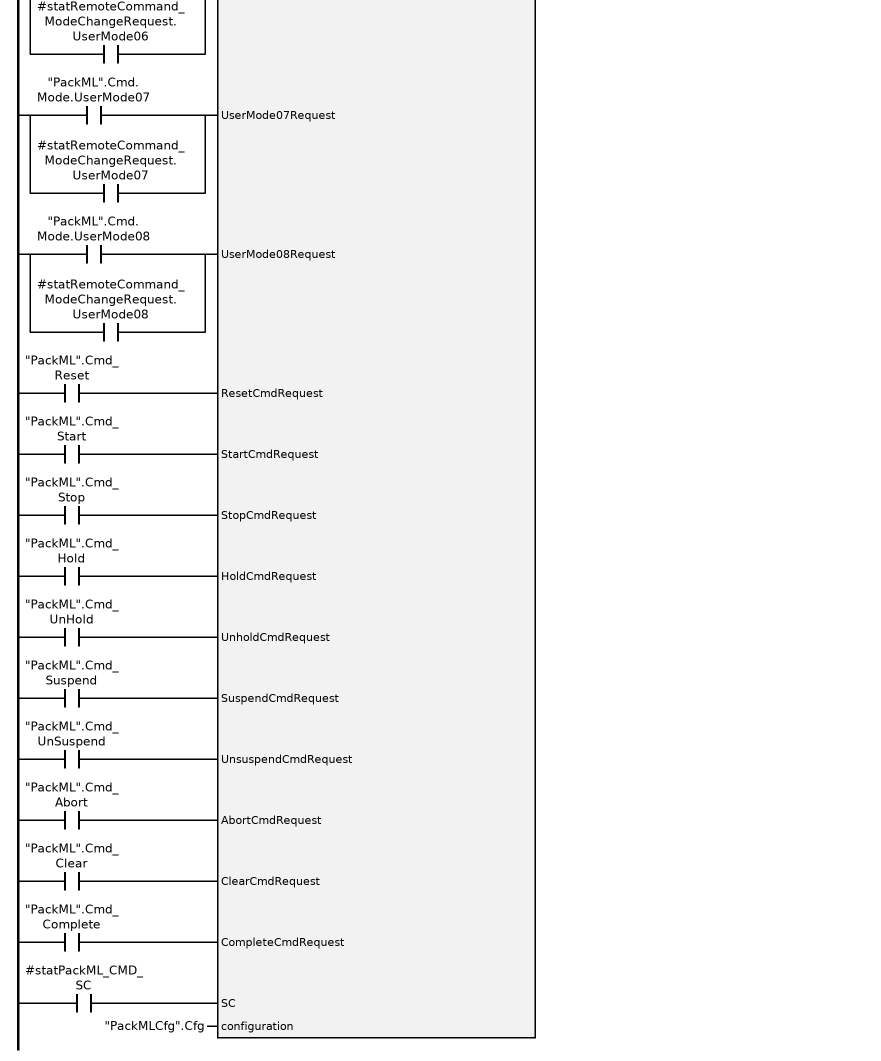
   RUNG wire#powerrail
      I_Contact( "FirstScan" )
      #instUnitModeStateManager(ProductionModeRequest := wire#w1, MaintenanceModeRequest := wire#w2, ManualModeRequest := wire#w3, UserMode01Request := wire#w4, UserMode02Request := wire#w5, UserMode03Request := wire#w6, UserMode04Request := wire#w7, UserMode05Request := wire#w8, UserMode06Request := wire#w9, UserMode07Request := wire#w10, UserMode08Request := wire#w11, ResetCmdRequest := wire#w12, StartCmdRequest := wire#w13, StopCmdRequest := wire#w14, HoldCmdRequest := wire#w15, UnholdCmdRequest := wire#w16, SuspendCmdRequest := wire#w17, UnsuspendCmdRequest := wire#w18, AbortCmdRequest := wire#w19, ClearCmdRequest := wire#w20, CompleteCmdRequest := wire#w21, SC := wire#w22, UnitMode :=, UnitModeChangeRequest := FALSE, CntrlCmd :=, CmdChangeRequest := FALSE, enableBooleanInterface := TRUE, configuration := "PackMLCfg".Cfg, UnitModeCurrent => "PackTags".Status.UnitModeCurrent, UnitModeRequested =>, UnitModeChangeInProcess => "PackTags".Status.UnitModeChangeInProcess, StateCurrent => "PackTags".Status.StateCurrent, StateRequested =>, StateChangeInProcess => "PackTags".Status.StateChangeInProcess, ProductionModeActive => "PackML".Sts.Mode.Production, MaintenanceModeActive => "PackML".Sts.Mode.Maintenance, ManualModeActive => "PackML".Sts.Mode.Manual, UserMode01Active => "PackML".Sts.Mode.UserMode01, UserMode02Active => "PackML".Sts.Mode.UserMode02, UserMode03Active => "PackML".Sts.Mode.UserMode03, UserMode04Active => "PackML".Sts.Mode.UserMode04, UserMode05Active => "PackML".Sts.Mode.UserMode05, UserMode06Active => "PackML".Sts.Mode.UserMode06, UserMode07Active => "PackML".Sts.Mode.UserMode07, UserMode08Active => "PackML".Sts.Mode.UserMode08, ClearingStateActive => "PackML".Sts.State.Clearing, StoppedStateActive => "PackML".Sts.State.Stopped, StartingStateActive => "PackML".Sts.State.Starting, IdleStateActive => "PackML".Sts.State.Idle, SuspendedStateActive => "PackML".Sts.State.Suspended, ExecuteStateActive => "PackML".Sts.State.Execute, StoppingStateActive => "PackML".Sts.State.Stopping, AbortingStateActive => "PackML".Sts.State.Aborting, AbortedStateActive => "PackML".Sts.State.Aborted, HoldingStateActive => "PackML".Sts.State.Holding, HeldStateActive => "PackML".Sts.State.Held, UnholdingStateActive => "PackML".Sts.State.Unholding, SuspendingStateActive => "PackML".Sts.State.Suspending, UnsuspendingStateActive => "PackML".Sts.State.Unsuspending, ResettingStateActive => "PackML".Sts.State.Resetting, CompletingStateActive => "PackML".Sts.State.Completing, CompleteStateActive => "PackML".Sts.State.Complete, StatesDisabled => "PackTags".Admin.StatesDisabled, diagnostics => "PackML".PackMLDiag)
      R_Coil( #statPackML_CMD_SC )
   END_RUNG
   RUNG wire#powerrail
      Contact( "PackML".Cmd.Mode.Production )
   END_RUNG wire#w1
   RUNG wire#powerrail
      Contact( #statRemoteCommand_ModeChangeRequest.Production )
   END_RUNG wire#w1
   RUNG wire#powerrail
      Contact( "PackML".Cmd.Mode.Maintenance )
   END_RUNG wire#w2
   RUNG wire#powerrail
      Contact( #statRemoteCommand_ModeChangeRequest.Maintenance )
   END_RUNG wire#w2
   RUNG wire#powerrail
      Contact( "PackML".Cmd.Mode.Manual )
   END_RUNG wire#w3
   RUNG wire#powerrail
      Contact( #statRemoteCommand_ModeChangeRequest.Manual )
   END_RUNG wire#w3
   RUNG wire#powerrail
      Contact( "PackML".Cmd.Mode.UserMode01 )
   END_RUNG wire#w4
   RUNG wire#powerrail
      Contact( #statRemoteCommand_ModeChangeRequest.UserMode01 )
   END_RUNG wire#w4
   RUNG wire#powerrail
      Contact( "PackML".Cmd.Mode.UserMode02 )
   END_RUNG wire#w5
   RUNG wire#powerrail
      Contact( #statRemoteCommand_ModeChangeRequest.UserMode02 )
   END_RUNG wire#w5
   RUNG wire#powerrail
      Contact( "PackML".Cmd.Mode.UserMode03 )
   END_RUNG wire#w6
   RUNG wire#powerrail
      Contact( #statRemoteCommand_ModeChangeRequest.UserMode03 )
   END_RUNG wire#w6
   RUNG wire#powerrail
      Contact( "PackML".Cmd.Mode.UserMode04 )
   END_RUNG wire#w7
   RUNG wire#powerrail
      Contact( #statRemoteCommand_ModeChangeRequest.UserMode04 )
   END_RUNG wire#w7
   RUNG wire#powerrail
      Contact( "PackML".Cmd.Mode.UserMode05 )
   END_RUNG wire#w8
   RUNG wire#powerrail
      Contact( #statRemoteCommand_ModeChangeRequest.UserMode05 )
   END_RUNG wire#w8
   RUNG wire#powerrail
      Contact( "PackML".Cmd.Mode.UserMode06 )
   END_RUNG wire#w9
   RUNG wire#powerrail
      Contact( #statRemoteCommand_ModeChangeRequest.UserMode06 )
   END_RUNG wire#w9
   RUNG wire#powerrail
      Contact( "PackML".Cmd.Mode.UserMode07 )
   END_RUNG wire#w10
   RUNG wire#powerrail
      Contact( #statRemoteCommand_ModeChangeRequest.UserMode07 )
   END_RUNG wire#w10
   RUNG wire#powerrail
      Contact( "PackML".Cmd.Mode.UserMode08 )
   END_RUNG wire#w11
   RUNG wire#powerrail
      Contact( #statRemoteCommand_ModeChangeRequest.UserMode08 )
   END_RUNG wire#w11
   RUNG wire#powerrail
      Contact( "PackML".Cmd_Reset )
   END_RUNG wire#w12
   RUNG wire#powerrail
      Contact( "PackML".Cmd_Start )
   END_RUNG wire#w13
   RUNG wire#powerrail
      Contact( "PackML".Cmd_Stop )
   END_RUNG wire#w14
   RUNG wire#powerrail
      Contact( "PackML".Cmd_Hold )
   END_RUNG wire#w15
   RUNG wire#powerrail
      Contact( "PackML".Cmd_UnHold )
   END_RUNG wire#w16
   RUNG wire#powerrail
      Contact( "PackML".Cmd_Suspend )
   END_RUNG wire#w17
   RUNG wire#powerrail
      Contact( "PackML".Cmd_UnSuspend )
   END_RUNG wire#w18
   RUNG wire#powerrail
      Contact( "PackML".Cmd_Abort )
   END_RUNG wire#w19
   RUNG wire#powerrail
      Contact( "PackML".Cmd_Clear )
   END_RUNG wire#w20
   RUNG wire#powerrail
      Contact( "PackML".Cmd_Complete )
   END_RUNG wire#w21
   RUNG wire#powerrail
      Contact( #statPackML_CMD_SC )
   END_RUNG wire#w22
   // the same network as SCL:
   #instUnitModeStateManager(EN := NOT "FirstScan",   // "LPMLV30_UnitModeStateManager"
                           UnitModeChangeRequest := FALSE,
                           CmdChangeRequest := FALSE,
                           enableBooleanInterface := TRUE,
                           ProductionModeRequest := "PackML".Cmd.Mode.Production OR #statRemoteCommand_ModeChangeRequest.Production,
                           MaintenanceModeRequest := "PackML".Cmd.Mode.Maintenance OR #statRemoteCommand_ModeChangeRequest.Maintenance,
                           ManualModeRequest := "PackML".Cmd.Mode.Manual OR #statRemoteCommand_ModeChangeRequest.Manual,
                           UserMode01Request := "PackML".Cmd.Mode.UserMode01 OR #statRemoteCommand_ModeChangeRequest.UserMode01,
                           UserMode02Request := "PackML".Cmd.Mode.UserMode02 OR #statRemoteCommand_ModeChangeRequest.UserMode02,
                           UserMode03Request := "PackML".Cmd.Mode.UserMode03 OR #statRemoteCommand_ModeChangeRequest.UserMode03,
                           UserMode04Request := "PackML".Cmd.Mode.UserMode04 OR #statRemoteCommand_ModeChangeRequest.UserMode04,
                           UserMode05Request := "PackML".Cmd.Mode.UserMode05 OR #statRemoteCommand_ModeChangeRequest.UserMode05,
                           UserMode06Request := "PackML".Cmd.Mode.UserMode06 OR #statRemoteCommand_ModeChangeRequest.UserMode06,
                           UserMode07Request := "PackML".Cmd.Mode.UserMode07 OR #statRemoteCommand_ModeChangeRequest.UserMode07,
                           UserMode08Request := "PackML".Cmd.Mode.UserMode08 OR #statRemoteCommand_ModeChangeRequest.UserMode08,
                           ResetCmdRequest := "PackML".Cmd_Reset,
                           StartCmdRequest := "PackML".Cmd_Start,
                           StopCmdRequest := "PackML".Cmd_Stop,
                           HoldCmdRequest := "PackML".Cmd_Hold,
                           UnholdCmdRequest := "PackML".Cmd_UnHold,
                           SuspendCmdRequest := "PackML".Cmd_Suspend,
                           UnsuspendCmdRequest := "PackML".Cmd_UnSuspend,
                           AbortCmdRequest := "PackML".Cmd_Abort,
                           ClearCmdRequest := "PackML".Cmd_Clear,
                           CompleteCmdRequest := "PackML".Cmd_Complete,
                           SC := #statPackML_CMD_SC,
                           configuration := "PackMLCfg".Cfg,
                           UnitModeCurrent => "PackTags".Status.UnitModeCurrent,
                           UnitModeChangeInProcess => "PackTags".Status.UnitModeChangeInProcess,
                           StateCurrent => "PackTags".Status.StateCurrent,
                           StateChangeInProcess => "PackTags".Status.StateChangeInProcess,
                           ProductionModeActive => "PackML".Sts.Mode.Production,
                           MaintenanceModeActive => "PackML".Sts.Mode.Maintenance,
                           ManualModeActive => "PackML".Sts.Mode.Manual,
                           UserMode01Active => "PackML".Sts.Mode.UserMode01,
                           UserMode02Active => "PackML".Sts.Mode.UserMode02,
                           UserMode03Active => "PackML".Sts.Mode.UserMode03,
                           UserMode04Active => "PackML".Sts.Mode.UserMode04,
                           UserMode05Active => "PackML".Sts.Mode.UserMode05,
                           UserMode06Active => "PackML".Sts.Mode.UserMode06,
                           UserMode07Active => "PackML".Sts.Mode.UserMode07,
                           UserMode08Active => "PackML".Sts.Mode.UserMode08,
                           ClearingStateActive => "PackML".Sts.State.Clearing,
                           StoppedStateActive => "PackML".Sts.State.Stopped,
                           StartingStateActive => "PackML".Sts.State.Starting,
                           IdleStateActive => "PackML".Sts.State.Idle,
                           SuspendedStateActive => "PackML".Sts.State.Suspended,
                           ExecuteStateActive => "PackML".Sts.State.Execute,
                           StoppingStateActive => "PackML".Sts.State.Stopping,
                           AbortingStateActive => "PackML".Sts.State.Aborting,
                           AbortedStateActive => "PackML".Sts.State.Aborted,
                           HoldingStateActive => "PackML".Sts.State.Holding,
                           HeldStateActive => "PackML".Sts.State.Held,
                           UnholdingStateActive => "PackML".Sts.State.Unholding,
                           SuspendingStateActive => "PackML".Sts.State.Suspending,
                           UnsuspendingStateActive => "PackML".Sts.State.Unsuspending,
                           ResettingStateActive => "PackML".Sts.State.Resetting,
                           CompletingStateActive => "PackML".Sts.State.Completing,
                           CompleteStateActive => "PackML".Sts.State.Complete,
                           StatesDisabled => "PackTags".Admin.StatesDisabled,
                           diagnostics => "PackML".PackMLDiag,
                           ENO => #_w1);
   IF #_w1 THEN #statPackML_CMD_SC := FALSE; END_IF;
END_REGION

REGION Network 15: "Times" used to format PackML.Admin times and for the HMI display
   // PackML State and Mode Times for HMI
   // 
   // The times spent in each mode and state are calculated in the PackML FB.  This 
   // FB is used to move the modes and states time arrays (current and cumulative 
   // times) into a single array - that is based upon the curent mode - for both 
   // current and cumlative state times.   This single arry is used by the HMI
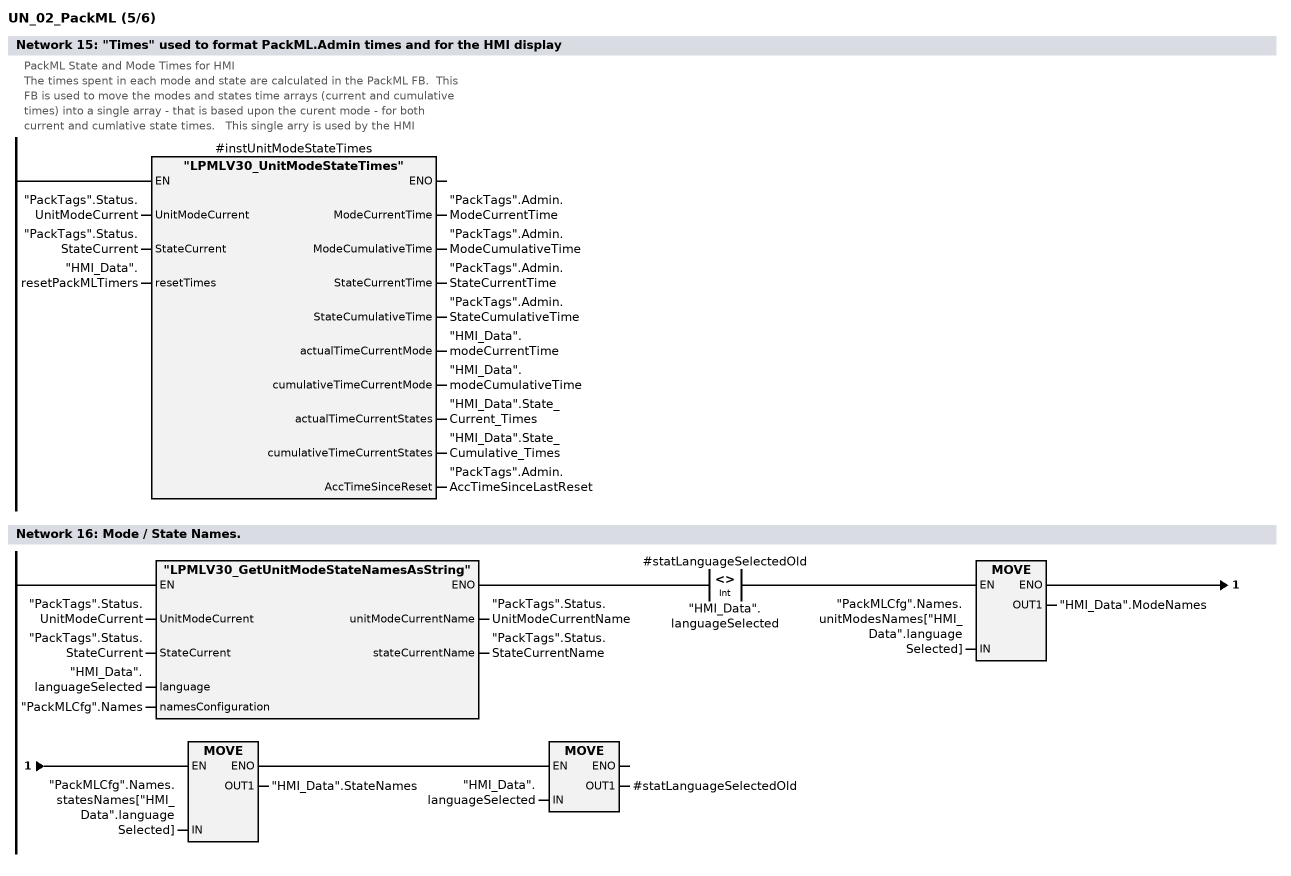
   RUNG wire#powerrail
      #instUnitModeStateTimes(UnitModeCurrent := "PackTags".Status.UnitModeCurrent, StateCurrent := "PackTags".Status.StateCurrent, resetTimes := "HMI_Data".resetPackMLTimers, ModeCurrentTime => "PackTags".Admin.ModeCurrentTime, ModeCumulativeTime => "PackTags".Admin.ModeCumulativeTime, StateCurrentTime => "PackTags".Admin.StateCurrentTime, StateCumulativeTime => "PackTags".Admin.StateCumulativeTime, actualTimeCurrentMode => "HMI_Data".modeCurrentTime, cumulativeTimeCurrentMode => "HMI_Data".modeCumulativeTime, actualTimeCurrentStates => "HMI_Data".State_Current_Times, cumulativeTimeCurrentStates => "HMI_Data".State_Cumulative_Times, AccTimeSinceReset => "PackTags".Admin.AccTimeSinceLastReset)
   END_RUNG
   // the same network as SCL:
   #instUnitModeStateTimes(UnitModeCurrent := "PackTags".Status.UnitModeCurrent,   // "LPMLV30_UnitModeStateTimes"
                           StateCurrent := "PackTags".Status.StateCurrent,
                           resetTimes := "HMI_Data".resetPackMLTimers,
                           ModeCurrentTime => "PackTags".Admin.ModeCurrentTime,
                           ModeCumulativeTime => "PackTags".Admin.ModeCumulativeTime,
                           StateCurrentTime => "PackTags".Admin.StateCurrentTime,
                           StateCumulativeTime => "PackTags".Admin.StateCumulativeTime,
                           actualTimeCurrentMode => "HMI_Data".modeCurrentTime,
                           cumulativeTimeCurrentMode => "HMI_Data".modeCumulativeTime,
                           actualTimeCurrentStates => "HMI_Data".State_Current_Times,
                           cumulativeTimeCurrentStates => "HMI_Data".State_Cumulative_Times,
                           AccTimeSinceReset => "PackTags".Admin.AccTimeSinceLastReset);
END_REGION

REGION Network 16: Mode / State Names.
   RUNG wire#powerrail
      "LPMLV30_GetUnitModeStateNamesAsString"(UnitModeCurrent := "PackTags".Status.UnitModeCurrent, StateCurrent := "PackTags".Status.StateCurrent, language := "HMI_Data".languageSelected, namesConfiguration := "PackMLCfg".Names, unitModeCurrentName => "PackTags".Status.UnitModeCurrentName, stateCurrentName => "PackTags".Status.StateCurrentName)
      { S7_Templates := "SrcType := Int" } NE_Contact(in1 := #statLanguageSelectedOld, in2 := "HMI_Data".languageSelected)
      Move(in := "PackMLCfg".Names.unitModesNames["HMI_Data".languageSelected], out1 => "HMI_Data".ModeNames)
      Move(in := "PackMLCfg".Names.statesNames["HMI_Data".languageSelected], out1 => "HMI_Data".StateNames)
      Move(in := "HMI_Data".languageSelected, out1 => #statLanguageSelectedOld)
   END_RUNG
   // the same network as SCL:
   "LPMLV30_GetUnitModeStateNamesAsString"(UnitModeCurrent := "PackTags".Status.UnitModeCurrent,
                           StateCurrent := "PackTags".Status.StateCurrent,
                           language := "HMI_Data".languageSelected,
                           namesConfiguration := "PackMLCfg".Names,
                           unitModeCurrentName => "PackTags".Status.UnitModeCurrentName,
                           stateCurrentName => "PackTags".Status.StateCurrentName,
                           ENO => #_w1);
   IF #_w1 AND (#statLanguageSelectedOld <> "HMI_Data".languageSelected) THEN
       "HMI_Data".ModeNames := "PackMLCfg".Names.unitModesNames["HMI_Data".languageSelected];
       "HMI_Data".StateNames := "PackMLCfg".Names.statesNames["HMI_Data".languageSelected];
       #statLanguageSelectedOld := "HMI_Data".languageSelected;
   END_IF;
END_REGION

REGION Network 17: State Complete Commands
END_REGION

REGION Network 18: Set the State Complete (SC) bit
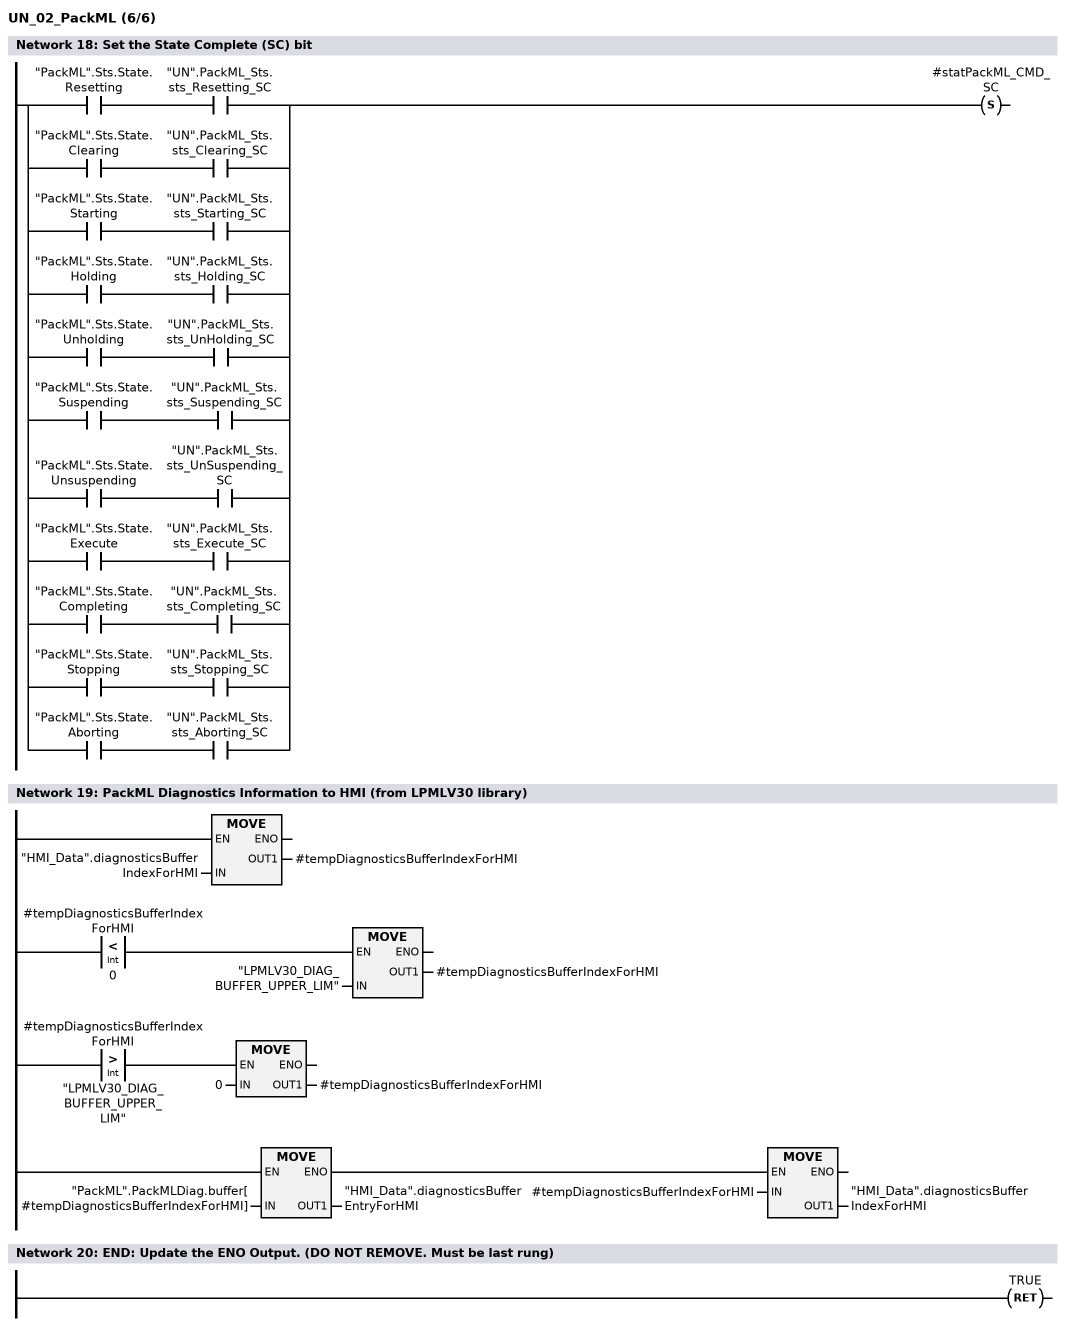
   RUNG wire#powerrail
      Contact( "PackML".Sts.State.Resetting )
      Contact( "UN".PackML_Sts.sts_Resetting_SC )
      wire#w1
      S_Coil( #statPackML_CMD_SC )
   END_RUNG
   RUNG wire#powerrail
      Contact( "PackML".Sts.State.Clearing )
      Contact( "UN".PackML_Sts.sts_Clearing_SC )
   END_RUNG wire#w1
   RUNG wire#powerrail
      Contact( "PackML".Sts.State.Starting )
      Contact( "UN".PackML_Sts.sts_Starting_SC )
   END_RUNG wire#w1
   RUNG wire#powerrail
      Contact( "PackML".Sts.State.Holding )
      Contact( "UN".PackML_Sts.sts_Holding_SC )
   END_RUNG wire#w1
   RUNG wire#powerrail
      Contact( "PackML".Sts.State.Unholding )
      Contact( "UN".PackML_Sts.sts_UnHolding_SC )
   END_RUNG wire#w1
   RUNG wire#powerrail
      Contact( "PackML".Sts.State.Suspending )
      Contact( "UN".PackML_Sts.sts_Suspending_SC )
   END_RUNG wire#w1
   RUNG wire#powerrail
      Contact( "PackML".Sts.State.Unsuspending )
      Contact( "UN".PackML_Sts.sts_UnSuspending_SC )
   END_RUNG wire#w1
   RUNG wire#powerrail
      Contact( "PackML".Sts.State.Execute )
      Contact( "UN".PackML_Sts.sts_Execute_SC )
   END_RUNG wire#w1
   RUNG wire#powerrail
      Contact( "PackML".Sts.State.Completing )
      Contact( "UN".PackML_Sts.sts_Completing_SC )
   END_RUNG wire#w1
   RUNG wire#powerrail
      Contact( "PackML".Sts.State.Stopping )
      Contact( "UN".PackML_Sts.sts_Stopping_SC )
   END_RUNG wire#w1
   RUNG wire#powerrail
      Contact( "PackML".Sts.State.Aborting )
      Contact( "UN".PackML_Sts.sts_Aborting_SC )
   END_RUNG wire#w1
   // the same network as SCL:
   IF ("PackML".Sts.State.Resetting AND "UN".PackML_Sts.sts_Resetting_SC) OR ("PackML".Sts.State.Clearing AND "UN".PackML_Sts.sts_Clearing_SC) OR ("PackML".Sts.State.Starting AND "UN".PackML_Sts.sts_Starting_SC) OR ("PackML".Sts.State.Holding AND "UN".PackML_Sts.sts_Holding_SC) OR ("PackML".Sts.State.Unholding AND "UN".PackML_Sts.sts_UnHolding_SC) OR ("PackML".Sts.State.Suspending AND "UN".PackML_Sts.sts_Suspending_SC) OR ("PackML".Sts.State.Unsuspending AND "UN".PackML_Sts.sts_UnSuspending_SC) OR ("PackML".Sts.State.Execute AND "UN".PackML_Sts.sts_Execute_SC) OR ("PackML".Sts.State.Completing AND "UN".PackML_Sts.sts_Completing_SC) OR ("PackML".Sts.State.Stopping AND "UN".PackML_Sts.sts_Stopping_SC) OR ("PackML".Sts.State.Aborting AND "UN".PackML_Sts.sts_Aborting_SC) THEN
       #statPackML_CMD_SC := TRUE;
   END_IF;
END_REGION

REGION Network 19: PackML Diagnostics Information to HMI (from LPMLV30 library)
   RUNG wire#powerrail
      Move(in := "HMI_Data".diagnosticsBufferIndexForHMI, out1 => #tempDiagnosticsBufferIndexForHMI)
   END_RUNG
   RUNG wire#powerrail
      { S7_Templates := "SrcType := Int" } LT_Contact(in1 := #tempDiagnosticsBufferIndexForHMI, in2 := 0)
      Move(in := "LPMLV30_DIAG_BUFFER_UPPER_LIM", out1 => #tempDiagnosticsBufferIndexForHMI)
   END_RUNG
   RUNG wire#powerrail
      { S7_Templates := "SrcType := Int" } GT_Contact(in1 := #tempDiagnosticsBufferIndexForHMI, in2 := "LPMLV30_DIAG_BUFFER_UPPER_LIM")
      Move(in := 0, out1 => #tempDiagnosticsBufferIndexForHMI)
   END_RUNG
   RUNG wire#powerrail
      Move(in := "PackML".PackMLDiag.buffer[#tempDiagnosticsBufferIndexForHMI], out1 => "HMI_Data".diagnosticsBufferEntryForHMI)
      Move(in := #tempDiagnosticsBufferIndexForHMI, out1 => "HMI_Data".diagnosticsBufferIndexForHMI)
   END_RUNG
   // the same network as SCL:
   #tempDiagnosticsBufferIndexForHMI := "HMI_Data".diagnosticsBufferIndexForHMI;
   IF #tempDiagnosticsBufferIndexForHMI < 0 THEN
       #tempDiagnosticsBufferIndexForHMI := "LPMLV30_DIAG_BUFFER_UPPER_LIM";
   END_IF;
   IF #tempDiagnosticsBufferIndexForHMI > "LPMLV30_DIAG_BUFFER_UPPER_LIM" THEN
       #tempDiagnosticsBufferIndexForHMI := 0;
   END_IF;
   "HMI_Data".diagnosticsBufferEntryForHMI := "PackML".PackMLDiag.buffer[#tempDiagnosticsBufferIndexForHMI];
   "HMI_Data".diagnosticsBufferIndexForHMI := #tempDiagnosticsBufferIndexForHMI;
END_REGION

REGION Network 20: END: Update the ENO Output. (DO NOT REMOVE. Must be last rung)
   RUNG wire#powerrail
      ReturnCoil( TRUE )
   END_RUNG
   // the same network as SCL:
   ENO := TRUE;
   RETURN;
END_REGION
END_FUNCTION_BLOCK

FUNCTION_BLOCK "UN_03_LineComm"   // FB31623, LAD
TITLE = UN_03_LineComm
{ S7_Optimized_Access := 'TRUE' }
AUTHOR : tech.team.motioncontrol@siemens.com
FAMILY : CPG
VERSION : 1.0
// Support: tech.team.motioncontrol@siemens.com
// Fax: +49 (0) 9131/98-1297
   VAR
      instAlarmRemoteStop : "CPG_Event";   // Remote Command - Stop
      instAlarmRemoteAbort : "CPG_Event";   // Remote Command - Abort
      instAlarmRemoteSuspendBlocked : "CPG_Event";   // Remote Command - Suspend (Blocked)
      instAlarmRemoteSuspendStarved : "CPG_Event";   // Remote Command - Suspend (Starved)
      instAlarmRemoteHold : "CPG_Event";   // Remote Command - Hold
      statRemoteSuspendCommand : Bool;   // Remote Suspend Command is active (from remote station)
      statRemoteHoldCommand : Bool;   // Remote Hold Command is active (from remote station)
   END_VAR
BEGIN

REGION Network 1: *** COMMUNICATION LOGIC ***
END_REGION

REGION Network 2: *** REMOTE COMMAND LOGIC ***
END_REGION

REGION Network 3: Remote Stop Command
   // "PackTags".Command.CntrlCmd = 3 (stop command value)
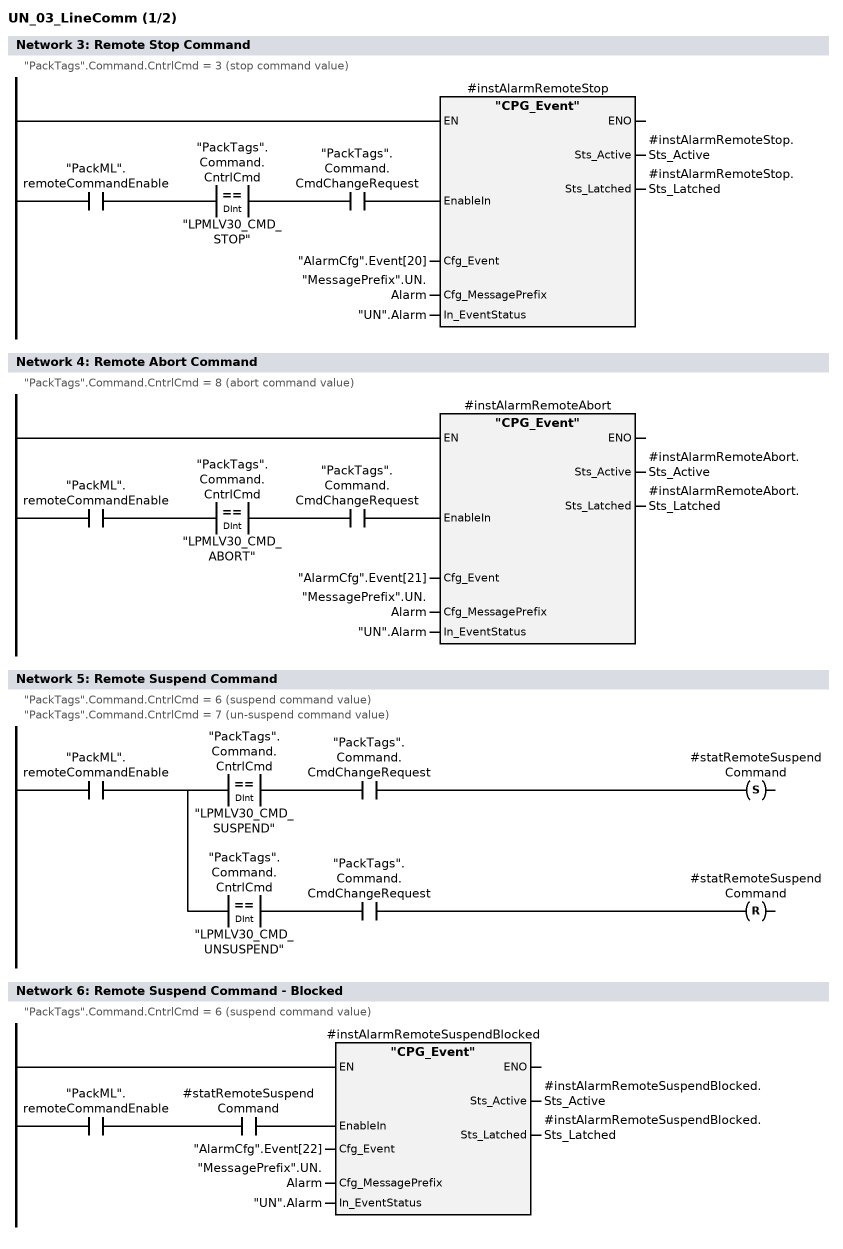
   RUNG wire#powerrail
      #instAlarmRemoteStop(EnableIn := wire#w1, Cfg_Event := "AlarmCfg".Event[20], Cfg_MessagePrefix := "MessagePrefix".UN.Alarm, In_EventStatus := "UN".Alarm, Sts_Active => #instAlarmRemoteStop.Sts_Active, Sts_Latched => #instAlarmRemoteStop.Sts_Latched)
   END_RUNG
   RUNG wire#powerrail
      Contact( "PackML".remoteCommandEnable )
      { S7_Templates := "SrcType := DInt" } EQ_Contact(in1 := "PackTags".Command.CntrlCmd, in2 := "LPMLV30_CMD_STOP")
      Contact( "PackTags".Command.CmdChangeRequest )
   END_RUNG wire#w1
   // the same network as SCL:
   #instAlarmRemoteStop(EnableIn := "PackML".remoteCommandEnable AND ("PackTags".Command.CntrlCmd = "LPMLV30_CMD_STOP") AND "PackTags".Command.CmdChangeRequest,   // "CPG_Event"
                        Cfg_Event := "AlarmCfg".Event[20],
                        Cfg_MessagePrefix := "MessagePrefix".UN.Alarm,
                        In_EventStatus := "UN".Alarm,
                        Sts_Active => #instAlarmRemoteStop.Sts_Active,
                        Sts_Latched => #instAlarmRemoteStop.Sts_Latched);
END_REGION

REGION Network 4: Remote Abort Command
   // "PackTags".Command.CntrlCmd = 8 (abort command value)
   RUNG wire#powerrail
      #instAlarmRemoteAbort(EnableIn := wire#w1, Cfg_Event := "AlarmCfg".Event[21], Cfg_MessagePrefix := "MessagePrefix".UN.Alarm, In_EventStatus := "UN".Alarm, Sts_Active => #instAlarmRemoteAbort.Sts_Active, Sts_Latched => #instAlarmRemoteAbort.Sts_Latched)
   END_RUNG
   RUNG wire#powerrail
      Contact( "PackML".remoteCommandEnable )
      { S7_Templates := "SrcType := DInt" } EQ_Contact(in1 := "PackTags".Command.CntrlCmd, in2 := "LPMLV30_CMD_ABORT")
      Contact( "PackTags".Command.CmdChangeRequest )
   END_RUNG wire#w1
   // the same network as SCL:
   #instAlarmRemoteAbort(EnableIn := "PackML".remoteCommandEnable AND ("PackTags".Command.CntrlCmd = "LPMLV30_CMD_ABORT") AND "PackTags".Command.CmdChangeRequest,   // "CPG_Event"
                         Cfg_Event := "AlarmCfg".Event[21],
                         Cfg_MessagePrefix := "MessagePrefix".UN.Alarm,
                         In_EventStatus := "UN".Alarm,
                         Sts_Active => #instAlarmRemoteAbort.Sts_Active,
                         Sts_Latched => #instAlarmRemoteAbort.Sts_Latched);
END_REGION

REGION Network 5: Remote Suspend Command
   // "PackTags".Command.CntrlCmd = 6 (suspend command value)
   // "PackTags".Command.CntrlCmd = 7 (un-suspend command value)
   RUNG wire#powerrail
      Contact( "PackML".remoteCommandEnable )
      wire#w1
      { S7_Templates := "SrcType := DInt" } EQ_Contact(in1 := "PackTags".Command.CntrlCmd, in2 := "LPMLV30_CMD_SUSPEND")
      Contact( "PackTags".Command.CmdChangeRequest )
      S_Coil( #statRemoteSuspendCommand )
   END_RUNG
   RUNG wire#w1
      { S7_Templates := "SrcType := DInt" } EQ_Contact(in1 := "PackTags".Command.CntrlCmd, in2 := "LPMLV30_CMD_UNSUSPEND")
      Contact( "PackTags".Command.CmdChangeRequest )
      R_Coil( #statRemoteSuspendCommand )
   END_RUNG
   // the same network as SCL:
   IF "PackML".remoteCommandEnable AND ("PackTags".Command.CntrlCmd = "LPMLV30_CMD_SUSPEND") AND "PackTags".Command.CmdChangeRequest THEN
       #statRemoteSuspendCommand := TRUE;
   END_IF;
   IF "PackML".remoteCommandEnable AND ("PackTags".Command.CntrlCmd = "LPMLV30_CMD_UNSUSPEND") AND "PackTags".Command.CmdChangeRequest THEN
       #statRemoteSuspendCommand := FALSE;
   END_IF;
END_REGION

REGION Network 6: Remote Suspend Command - Blocked
   // "PackTags".Command.CntrlCmd = 6 (suspend command value)
   RUNG wire#powerrail
      #instAlarmRemoteSuspendBlocked(EnableIn := wire#w1, Cfg_Event := "AlarmCfg".Event[22], Cfg_MessagePrefix := "MessagePrefix".UN.Alarm, In_EventStatus := "UN".Alarm, Sts_Active => #instAlarmRemoteSuspendBlocked.Sts_Active, Sts_Latched => #instAlarmRemoteSuspendBlocked.Sts_Latched)
   END_RUNG
   RUNG wire#powerrail
      Contact( "PackML".remoteCommandEnable )
      Contact( #statRemoteSuspendCommand )
   END_RUNG wire#w1
   // the same network as SCL:
   #instAlarmRemoteSuspendBlocked(EnableIn := "PackML".remoteCommandEnable AND #statRemoteSuspendCommand,   // "CPG_Event"
                           Cfg_Event := "AlarmCfg".Event[22],
                           Cfg_MessagePrefix := "MessagePrefix".UN.Alarm,
                           In_EventStatus := "UN".Alarm,
                           Sts_Active => #instAlarmRemoteSuspendBlocked.Sts_Active,
                           Sts_Latched => #instAlarmRemoteSuspendBlocked.Sts_Latched);
END_REGION

REGION Network 7: Remote Suspend Command - Starved
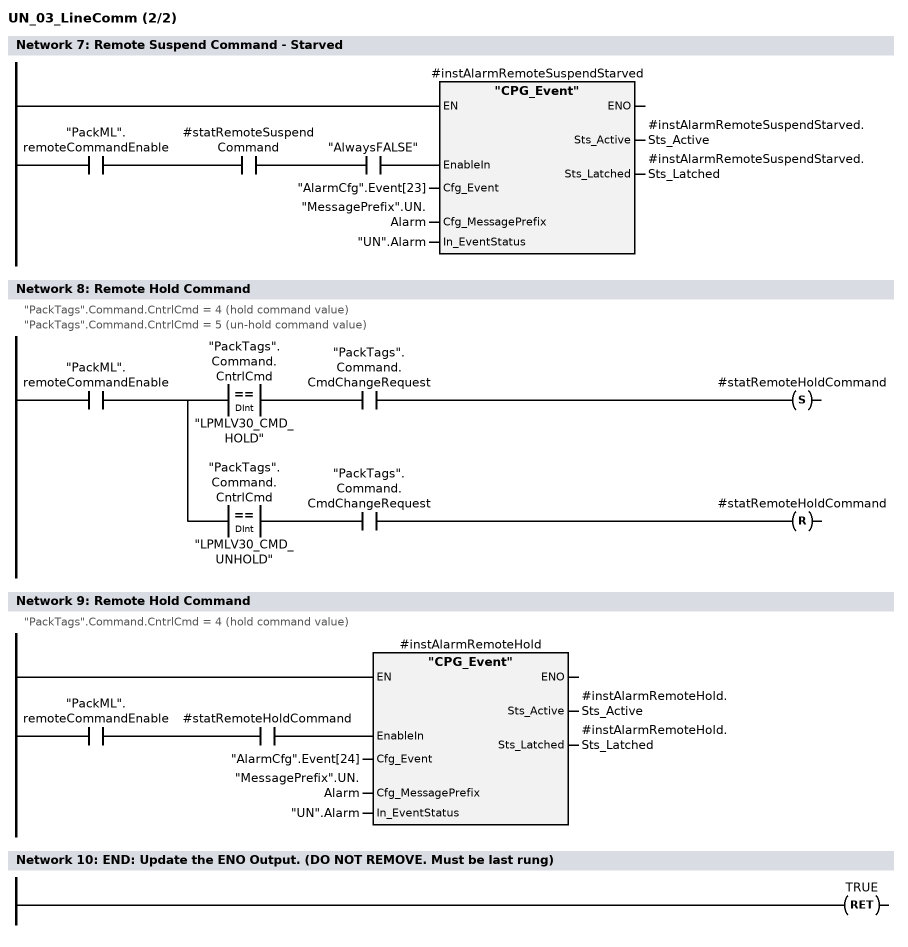
   RUNG wire#powerrail
      #instAlarmRemoteSuspendStarved(EnableIn := wire#w1, Cfg_Event := "AlarmCfg".Event[23], Cfg_MessagePrefix := "MessagePrefix".UN.Alarm, In_EventStatus := "UN".Alarm, Sts_Active => #instAlarmRemoteSuspendStarved.Sts_Active, Sts_Latched => #instAlarmRemoteSuspendStarved.Sts_Latched)
   END_RUNG
   RUNG wire#powerrail
      Contact( "PackML".remoteCommandEnable )
      Contact( #statRemoteSuspendCommand )
      Contact( "AlwaysFALSE" )
   END_RUNG wire#w1
   // the same network as SCL:
   #instAlarmRemoteSuspendStarved(EnableIn := "PackML".remoteCommandEnable AND #statRemoteSuspendCommand AND "AlwaysFALSE",   // "CPG_Event"
                           Cfg_Event := "AlarmCfg".Event[23],
                           Cfg_MessagePrefix := "MessagePrefix".UN.Alarm,
                           In_EventStatus := "UN".Alarm,
                           Sts_Active => #instAlarmRemoteSuspendStarved.Sts_Active,
                           Sts_Latched => #instAlarmRemoteSuspendStarved.Sts_Latched);
END_REGION

REGION Network 8: Remote Hold Command
   // "PackTags".Command.CntrlCmd = 4 (hold command value)
   // "PackTags".Command.CntrlCmd = 5 (un-hold command value)
   RUNG wire#powerrail
      Contact( "PackML".remoteCommandEnable )
      wire#w1
      { S7_Templates := "SrcType := DInt" } EQ_Contact(in1 := "PackTags".Command.CntrlCmd, in2 := "LPMLV30_CMD_HOLD")
      Contact( "PackTags".Command.CmdChangeRequest )
      S_Coil( #statRemoteHoldCommand )
   END_RUNG
   RUNG wire#w1
      { S7_Templates := "SrcType := DInt" } EQ_Contact(in1 := "PackTags".Command.CntrlCmd, in2 := "LPMLV30_CMD_UNHOLD")
      Contact( "PackTags".Command.CmdChangeRequest )
      R_Coil( #statRemoteHoldCommand )
   END_RUNG
   // the same network as SCL:
   IF "PackML".remoteCommandEnable AND ("PackTags".Command.CntrlCmd = "LPMLV30_CMD_HOLD") AND "PackTags".Command.CmdChangeRequest THEN
       #statRemoteHoldCommand := TRUE;
   END_IF;
   IF "PackML".remoteCommandEnable AND ("PackTags".Command.CntrlCmd = "LPMLV30_CMD_UNHOLD") AND "PackTags".Command.CmdChangeRequest THEN
       #statRemoteHoldCommand := FALSE;
   END_IF;
END_REGION

REGION Network 9: Remote Hold Command
   // "PackTags".Command.CntrlCmd = 4 (hold command value)
   RUNG wire#powerrail
      #instAlarmRemoteHold(EnableIn := wire#w1, Cfg_Event := "AlarmCfg".Event[24], Cfg_MessagePrefix := "MessagePrefix".UN.Alarm, In_EventStatus := "UN".Alarm, Sts_Active => #instAlarmRemoteHold.Sts_Active, Sts_Latched => #instAlarmRemoteHold.Sts_Latched)
   END_RUNG
   RUNG wire#powerrail
      Contact( "PackML".remoteCommandEnable )
      Contact( #statRemoteHoldCommand )
   END_RUNG wire#w1
   // the same network as SCL:
   #instAlarmRemoteHold(EnableIn := "PackML".remoteCommandEnable AND #statRemoteHoldCommand,   // "CPG_Event"
                        Cfg_Event := "AlarmCfg".Event[24],
                        Cfg_MessagePrefix := "MessagePrefix".UN.Alarm,
                        In_EventStatus := "UN".Alarm,
                        Sts_Active => #instAlarmRemoteHold.Sts_Active,
                        Sts_Latched => #instAlarmRemoteHold.Sts_Latched);
END_REGION

REGION Network 10: END: Update the ENO Output. (DO NOT REMOVE. Must be last rung)
   RUNG wire#powerrail
      ReturnCoil( TRUE )
   END_RUNG
   // the same network as SCL:
   ENO := TRUE;
   RETURN;
END_REGION
END_FUNCTION_BLOCK

FUNCTION_BLOCK "UN_04_EventControl"   // FB31624, LAD
TITLE = UN_04_EventControl
{ S7_Optimized_Access := 'TRUE' }
AUTHOR : tech.team.motioncontrol@siemens.com
FAMILY : CPG
VERSION : 1.1
// Support: tech.team.motioncontrol@siemens.com
   VAR
      instEventMgrAlarm : "CPG_EventManager";   // instance FB - Event Manager - Alarms Events
      instEventMgrWarning : "CPG_EventManager";   // instance FB - Event Manager - Warning Events
      instEventMgrStatus : "CPG_EventManager";   // instance FB - Event Manager - Status Events
      instStatusAlarmsNotReset : "CPG_Event";   // Status = Alarms Not Reset
      statEventMgr_Cmd_Reset : Bool;   // Reset Cmd for event managers
      statEventMgr_Cmd_Clear1stFlt : Bool;   // Clear 1st Fault Cmd for event managers
      statEventMgr_Clear1stFlt_OS : Bool;   // Clear 1st Fault Cmd - One shot
   END_VAR
   VAR_TEMP   // added for the SCL form of the ladder/FBD networks
      _w1 : Bool;
      _w2 : Bool;
   END_VAR
BEGIN

REGION Network 2: ** STATE MODEL REPORTING STATUS ****
END_REGION

REGION Network 3: *** Call the PackML Module Initialize Logic ***
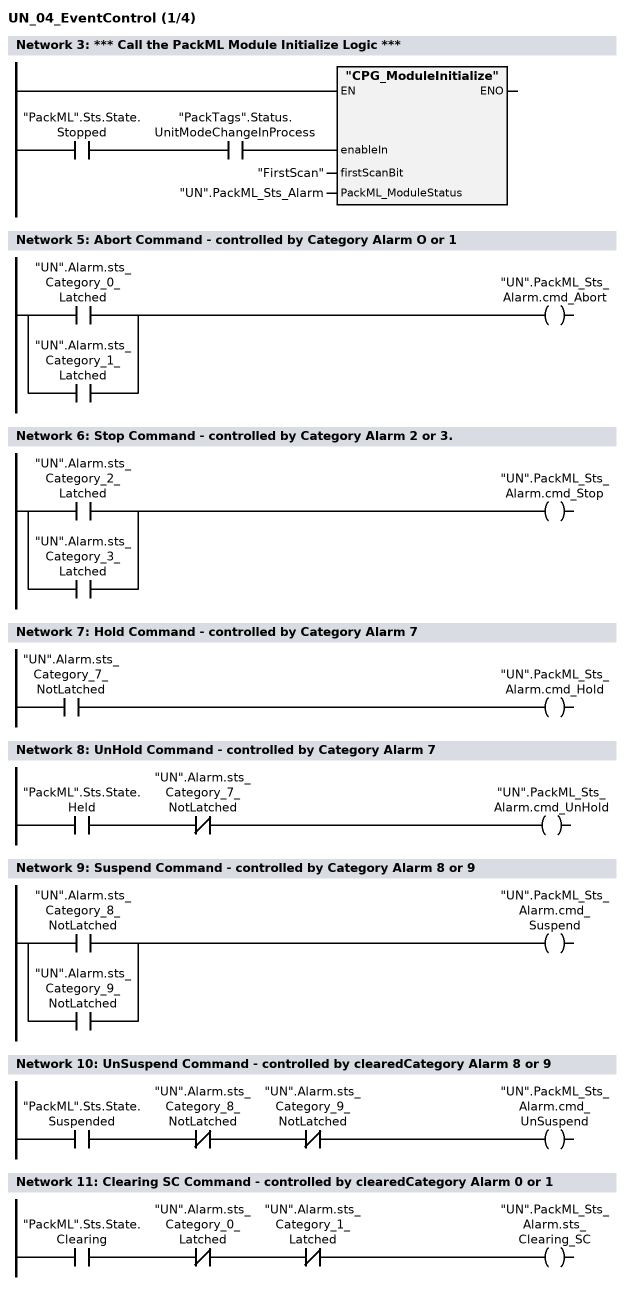
   RUNG wire#powerrail
      "CPG_ModuleInitialize"(enableIn := wire#w1, firstScanBit := "FirstScan", PackML_ModuleStatus := "UN".PackML_Sts_Alarm)
   END_RUNG
   RUNG wire#powerrail
      Contact( "PackML".Sts.State.Stopped )
      Contact( "PackTags".Status.UnitModeChangeInProcess )
   END_RUNG wire#w1
   // the same network as SCL:
   "CPG_ModuleInitialize"(enableIn := "PackML".Sts.State.Stopped AND "PackTags".Status.UnitModeChangeInProcess,
                          firstScanBit := "FirstScan",
                          PackML_ModuleStatus := "UN".PackML_Sts_Alarm);
END_REGION

REGION Network 4: Begin the LOGIC section.
END_REGION

REGION Network 5: Abort Command - controlled by Category Alarm O or 1
   RUNG wire#powerrail
      Contact( "UN".Alarm.sts_Category_0_Latched )
      wire#w1
      Coil( "UN".PackML_Sts_Alarm.cmd_Abort )
   END_RUNG
   RUNG wire#powerrail
      Contact( "UN".Alarm.sts_Category_1_Latched )
   END_RUNG wire#w1
   // the same network as SCL:
   "UN".PackML_Sts_Alarm.cmd_Abort := "UN".Alarm.sts_Category_0_Latched OR "UN".Alarm.sts_Category_1_Latched;
END_REGION

REGION Network 6: Stop Command - controlled by Category Alarm 2 or 3.
   RUNG wire#powerrail
      Contact( "UN".Alarm.sts_Category_2_Latched )
      wire#w1
      Coil( "UN".PackML_Sts_Alarm.cmd_Stop )
   END_RUNG
   RUNG wire#powerrail
      Contact( "UN".Alarm.sts_Category_3_Latched )
   END_RUNG wire#w1
   // the same network as SCL:
   "UN".PackML_Sts_Alarm.cmd_Stop := "UN".Alarm.sts_Category_2_Latched OR "UN".Alarm.sts_Category_3_Latched;
END_REGION

REGION Network 7: Hold Command - controlled by Category Alarm 7
   RUNG wire#powerrail
      Contact( "UN".Alarm.sts_Category_7_NotLatched )
      Coil( "UN".PackML_Sts_Alarm.cmd_Hold )
   END_RUNG
   // the same network as SCL:
   "UN".PackML_Sts_Alarm.cmd_Hold := "UN".Alarm.sts_Category_7_NotLatched;
END_REGION

